// TIA Portal project "Projekt_Serhii_Bodnia" (V19) (continued)

   REGION Timer
       #TP_Remover(IN:= #FlOp_Neg_LS_Auslauf_Band_1.Q,
                   PT:=T#500ms);
       // Störungserkennung: wenn LS_Auslauf länger als 3s aktiv und Band läuft → Stau
       #TON_Störung_LS_Einlauf_Band_0(IN := #LS_Einlauf_Band_0 AND #M_Band_0,
                            PT := T#3s);
       #TON_Störung_LS_Auslauf_Band_0(IN := #LS_Auslauf_Band_0 AND #M_Band_0,
                            PT := T#3s);
       #TON_Störung_LS_Einlauf_Band_1(IN := #LS_Einlauf_Band_1 AND #M_Band_1,
                            PT := T#3s);
       #TON_Störung_LS_Auslauf_Band_1 (IN := #LS_Auslauf_Band_1 AND #M_Band_1,
                            PT := T#3s);
       #TON_Störung_LS_Vision_Sensor (IN := #LS_Vision_Sensor AND #M_Band_0,
                            PT := T#3s);
       #TON_Störung_LS_Arm_0 (IN := #LS_Arm_0 AND #M_Band_0,
                            PT := T#3s);

   END_REGION

    REGION Produktarten
    // Produktart-Rezeptur-Mapping: HMI-Produktauswahl auf Farbewert umrechnen
       IF #Produktart_Linie_0 = 4 THEN
           #Rezeptur_Art_0 := 5;
       ELSIF #Produktart_Linie_0 = 2 THEN
           #Rezeptur_Art_0 := 6;
       END_IF;
       IF #Produktart_Linie_1 = 1 THEN
           #Rezeptur_Art_1 := 2;
       ELSIF #Produktart_Linie_1 = 2 THEN
           #Rezeptur_Art_1 := 1;
       END_IF;
   END_REGION

   REGION Meldungen
       // Störungserkennung: wenn LS_Einlauf oder LS_Auslauf länger als 3s aktiv und Band läuft → Stau
       IF ((#Teil_auf_Band_0 > 5 OR #TON_Störung_LS_Einlauf_Band_0.Q OR #TON_Störung_LS_Auslauf_Band_0.Q
           OR #TON_Störung_LS_Vision_Sensor.Q OR #TON_Störung_LS_Arm_0.Q) AND #M_Band_0 AND NOT #Stop_Modus)
           OR ((#Teil_auf_Band_1 > 5 OR #TON_Störung_LS_Einlauf_Band_1.Q OR #TON_Störung_LS_Auslauf_Band_1.Q) AND #M_Band_1 AND NOT #Stop_Modus) THEN
           // Störungsmerker setzen
           #M_Störung := TRUE;
       END_IF;
       // Störung über HMI quittieren: Bit des Quittierungswortes (HMI_Quittierung)
       IF #Quittierung THEN
           #M_Störung := FALSE;
       END_IF;


   END_REGION

   REGION Sortierung
       IF #FlOp_Pos_LS_Arm_0.Q THEN
           //Farbe des ersten  Werkstücks in der Warteschlange prüfen 
           #Current_Art := #Buffer[0];
           // Array verschieben
           FOR #i := 0 TO 4 DO
               #Buffer[#i] := #Buffer[#i + 1];
           END_FOR;
           // Letzten Element nach dem Verschiebung löschen und den Zäler verringern
           #Buffer[5] := 0;
           IF #Count > 0 THEN
               #Count := #Count - 1;
           END_IF;
       END_IF;

       // Ein- und Ausschaltung Arm_0
       IF #Start_Modus AND (#Current_Art = #Rezeptur_Art_0 AND #FlOp_Pos_LS_Arm_0.Q) THEN
           // Sortierarm EIN: wenn erkannte Produktart dem Rezept entspricht
           #M_Arm_turn_0 := TRUE;
           #M_Arm_Band_0 := TRUE;
       END_IF;
       IF #"FlOp_Neg_LS_Auslauf_Band_0 (1)".Q THEN
           // Arm ausschalten: wenn Teil den Auslauf Band 0 verlassen hat
           #M_Arm_turn_0 := FALSE;
           #M_Arm_Band_0 := FALSE;
       END_IF;

   END_REGION

   REGION Eintag in den Puffer

       IF #FlOp_Pos_LS_Vision_Sensor.Q THEN
           // Farbe speichern
           #Buffer[#Count] := #Vision_Sensor;
           // Platz für den nächsten vorbereiten
           #Count := #Count + 1;
       END_IF;
   END_REGION

   REGION Bänder
       REGION Band_0
           REGION Erfassung der Anzahl der Teileauf dem Band_0
               IF #Start_Modus AND NOT #Stop_Modus THEN
                   // Teilezähler Band_0: zählt aktuell transportierte Teile
                   IF #FlOp_Neg_LS_Einlauf_Band_0.Q THEN
                       #Teil_auf_Band_0 := #Teil_auf_Band_0 + 1;
                   END_IF;
                   IF #Teil_auf_Band_0 > 0 AND (#"FlOp_Neg_LS_Auslauf_Band_0 (1)".Q OR #"FlOp_Neg_LS_Auslauf_Band_0 (2)".Q) THEN
                       #Teil_auf_Band_0 := #Teil_auf_Band_0 - 1;
                   END_IF;
               END_IF;
               IF #Not_Aus_Modus OR #M_Störung THEN
                   #Teil_auf_Band_0 := 0;
               END_IF;
           END_REGION
           REGION Band_0 Steuerung
               // Band_0 läuft solange Teile vorhanden oder neu eingetroffen
               IF #Start_Modus AND (#FlOp_Neg_LS_Einlauf_Band_0.Q OR #Teil_auf_Band_0 > 0) THEN
                   #M_Band_0 := True;
               ELSE
                   #M_Band_0 := FALSE;
               END_IF;

           END_REGION
       END_REGION
       REGION Band_1
           REGION Erfassung der Anzahl der Teileauf dem Band_1
               IF #Start_Modus AND NOT #Stop_Modus THEN
                   // Teilezähler Band 1: zählt aktuell transportierte Teile
                   IF #FlOp_Pos_LS_Einlauf_Band_1.Q THEN
                       #Teil_auf_Band_1 := #Teil_auf_Band_1 + 1;
                   END_IF;
                   IF #Teil_auf_Band_1 > 0 AND #FlOp_Neg_LS_Auslauf_Band_1.Q THEN
                       #Teil_auf_Band_1 := #Teil_auf_Band_1 - 1;
                   END_IF;
               END_IF;
               IF #Not_Aus_Modus OR #M_Störung THEN
                   #Teil_auf_Band_1 := 0;
               END_IF;

           END_REGION
           REGION Band_1 Steuerung
               // Band_1 läuft solange Teile vorhanden oder neu eingetroffen
               IF #Start_Modus AND #FlOp_Pos_LS_Einlauf_Band_1.Q OR #Teil_auf_Band_1 > 0 THEN
                   #M_Band_1 := True;
               ELSE
                   #M_Band_1 := FALSE;
              END_IF;
           END_REGION

       END_REGION

   END_REGION

   REGION Actoren
       // Physische Ausgaben: Bänder und Sortierarm (gesperrt bei Stopp-Modus)
       #Band_0 := #M_Band_0 AND NOT #Stop_Modus;
       #Band_1 := #M_Band_1 AND NOT #Stop_Modus;
       #Arm_turn_0 := #M_Arm_turn_0 AND NOT #Stop_Modus;
       #Arm_Band_0 := #M_Arm_Band_0 AND NOT #Stop_Modus;
       #Remover := #TP_Remover.Q;
       // Gesamtanzahl Fertigteile für HMI
       #Anzahl_Kanister := #CTU_Kanister.CV;
       //
       #Störung := #M_Störung;
   END_REGION
END_FUNCTION_BLOCK

FUNCTION_BLOCK "FB_AbfüllmaschineBand_SCL"   // FB7, SCL
{ S7_Optimized_Access := 'TRUE' }
VERSION : 0.1
   VAR_INPUT
      Start_Mode : Bool;
      Stop_Mode : Bool;
      NotAus_Mode : Bool;
      LS_Einlauf : Bool;
      LS_Auslauf : Bool;
      Diff_Sensor_Tank : Bool;
      Dosing_Aktive : Bool;
      Tank_Level_Meter : Real;
      Quittierung : Bool;
   END_VAR
   VAR_OUTPUT
      Einlaufband : Bool;
      Start_Dosierung : Bool;
      Emitter : Bool;
      "Start Button (Light)" : Bool;
      "Stop Button (Light)" : Bool;
      "Stack Light (Green)" : Bool;
      "Stack Light (Red)" : Bool;
      "Stack Light (Yellow)" : Bool;
      Störung : Bool;
   END_VAR
   VAR
      Stat_Trigger_Neg_Dosing_Stand : F_TRIG;
      Stat_Trigger_Neg_LS_Auslauf : F_TRIG;
      TON_weit_500ms : TON_TIME;
      TON_Störung_Einlauf : TON_TIME;
      TON_Störung_Auslauf : TON_TIME;
      TON_Störung_LS_Tank : TON_TIME;
      iSchritt : Int;
      M_Einlaufband : Bool;
      M_Störung : Bool;
   END_VAR
BEGIN

   REGION Flankenabfragen
       // Statement section REGION
       #Stat_Trigger_Neg_Dosing_Stand(CLK := #Dosing_Aktive); // Fallende Flanke: Dosierung beendet
       #Stat_Trigger_Neg_LS_Auslauf(CLK := #LS_Auslauf); // Fallende Flanke: Flasche am Auslauf
   END_REGION

   REGION Timer
       // Störungserkennung: wenn LS_Einlauf oder LS_Auslauf oder LS_Tank länger als 10s aktiv und Band läuft → Stau
       #"TON_Störung_Einlauf"(IN := #LS_Einlauf AND #M_Einlaufband AND NOT #Stop_Mode,
                            PT := T#10s);
     #TON_Störung_Auslauf(IN := #LS_Auslauf AND #M_Einlaufband AND NOT #Stop_Mode,
                            PT := T#10s);
       #TON_Störung_LS_Tank(IN := #Diff_Sensor_Tank AND #M_Einlaufband AND NOT #Stop_Mode,
                            PT := T#10s);
   END_REGION


   REGION Meldungen
       // Störungserkennung: wenn LS_Einlauf oder LS_Auslauf oder LS_Tank länger als 10s aktiv und Band läuft → Stau

       IF #TON_Störung_Einlauf.Q OR #TON_Störung_Auslauf.Q OR #TON_Störung_LS_Tank.Q THEN
           // Störungsmerker setzen
           #M_Störung := TRUE;
       END_IF;
       // Störung über HMI quittieren: Bit des Quittierungswortes (HMI_Quittierung)
       IF #Quittierung THEN
           #M_Störung := FALSE;
       END_IF;

   END_REGION

   REGION Schrittkette
       IF #NotAus_Mode OR #M_Störung THEN
           // Not-Aus: sofortiger Rücksprung in Initialschritt (alle Aktoren werden abgeschaltet)
           #iSchritt := 0;
       END_IF;

       CASE #iSchritt OF
           0:  // Initialschritt: Startbedingungen prüfen
               // Start nur wenn: Startmodus aktiv UND Füllventil geschlossen UND Tank nicht leer
               IF #Start_Mode  AND (#Tank_Level_Meter >= 1) THEN
                   #iSchritt := 1;
               END_IF;
           1: // Emitter EIN: leere Kanister ausgeben; warten bis Kanister erkannt
               IF #LS_Einlauf THEN
                   #iSchritt := 2;
               END_IF;
           2: // Einlaufband EIN: Kanister unter den Dosierkopf transportieren
              // Übergang wenn Diffusionssensor der Kanister unter dem Tank detektiert
               IF #Diff_Sensor_Tank THEN
                   #iSchritt := 3;
               END_IF;
           3: // Einlaufband AUS; Dosierung starten; warten auf fallende Flanke (Dosierung beendet)
               IF #Stat_Trigger_Neg_Dosing_Stand.Q THEN
                   #iSchritt := 4;
               END_IF;
           4: // Einlaufband EIN (mit TON-Nachlauf 500ms): gefüllte Flasche zum Auslauf schieben
              // Übergang bei fallender Flanke: Kanister hat Auslaufsensor verlassen
               IF #Stat_Trigger_Neg_LS_Auslauf.Q THEN
                   #iSchritt := 1;
               END_IF;

           ELSE  // Unbekannter Schritt: Sicherheitshalber Rücksprung
               #iSchritt := 0;
       END_CASE;
   END_REGION
   REGION Actoren
      // 1. Emitter
       #Emitter := (#iSchritt = 1);
       // 2. Einlaufband
       #TON_weit_500ms(IN := (#iSchritt = 4), PT := T#500ms);
       #Einlaufband := ((#iSchritt = 2) OR #TON_weit_500ms.Q) AND NOT #Stop_Mode;
       #M_Einlaufband := ((#iSchritt = 2) OR #TON_weit_500ms.Q) AND NOT #Stop_Mode;
       // 3. Start_Dosierung
       #Start_Dosierung := (#iSchritt = 3) AND NOT #Stop_Mode;
       // 4. Signallleuchten
       #"Start Button (Light)" := #Start_Mode AND NOT #Stop_Mode;
       #"Stack Light (Green)" := #Start_Mode AND NOT #Stop_Mode;
       #"Stop Button (Light)" := #Stop_Mode;
       #"Stack Light (Red)" := #Stop_Mode;
       #"Stack Light (Yellow)" := #NotAus_Mode;
       //
       #Störung := #M_Störung;

   END_REGION
END_FUNCTION_BLOCK

FUNCTION_BLOCK "FB_Band mit Positionierleisten"   // FB8, SCL
{ S7_Optimized_Access := 'TRUE' }
VERSION : 0.1
   VAR_INPUT
      LS_Einlauf : Bool;
      LS_Auslauf : Bool;
      LS_Positionierer : Bool;
      Start_Modus : Bool;
      Stop_Modus : Bool;
      Not_Aus_Modus : Bool;
      Acknowledge : Bool;
      Quittierung : Bool;
   END_VAR
   VAR_OUTPUT
      Band : Bool;
      Positionierer : Bool;
      Ready_To_Send_Teil : Bool;
      Ready_To_Receive_Teil : Bool;
      Störung : Bool;
   END_VAR
   VAR
      FlOp_Pos_LS_Einlauf : R_TRIG;
      FlOp_Neg_LS_Einlauf : F_TRIG;
      FlOp_Neg_LS_Auslauf : F_TRIG;
      Teil_auf_Band : Int;
      M_Band : Bool;
      M_Positionierer : Bool;
      M_Störung : Bool;
      TON_Störung_LS_Einlauf : TON_TIME;
      TON_Störung_LS_Auslauf : TON_TIME;
      TON_Störung_LS_Positionierer : TON_TIME;
   END_VAR
BEGIN
   REGION Flankenabfragen
       // Alle Flanken müssen am Anfang des Bausteins ausgewertet werden
       #FlOp_Pos_LS_Einlauf(CLK := #LS_Einlauf);
       #FlOp_Neg_LS_Einlauf(CLK := #LS_Einlauf);
       #FlOp_Neg_LS_Auslauf(CLK := #LS_Auslauf);
   END_REGION

   REGION Timers
       // Störungserkennung: wenn LS_Einlauf oder LS_Auslauf länger als 10s aktiv und Band läuft → Stau
       #TON_Störung_LS_Einlauf(IN := #LS_Einlauf AND #M_Band AND NOT #Stop_Modus,
                               PT := T#10s);
       #TON_Störung_LS_Auslauf(IN := #LS_Auslauf AND #M_Band AND NOT #Stop_Modus,
                               PT := T#10s);
       #TON_Störung_LS_Positionierer (IN := #LS_Positionierer AND #M_Band AND NOT #Stop_Modus,
                               PT := T#10s);
   END_REGION

   REGION Meldungen
       // Störungserkennung: wenn LS_Einlauf oder LS_Auslauf länger als 10s aktiv und Band läuft → Stau
       IF #Teil_auf_Band > 3 OR #TON_Störung_LS_Einlauf.Q OR #TON_Störung_LS_Auslauf.Q OR #TON_Störung_LS_Positionierer.Q THEN
           // Störungsmerker setzen
           #M_Störung := TRUE;
       END_IF;
       // Störung über HMI quittieren: Bit des Quittierungswortes (HMI_Quittierung)
       IF #Quittierung THEN
           #M_Störung := FALSE;
       END_IF;

   END_REGION

   REGION Band
       // Teilezähler: zählt Teile auf dem Band
       IF #Start_Modus AND #FlOp_Neg_LS_Einlauf.Q THEN
           // Neues Teil aufgenommen
           #Teil_auf_Band := #Teil_auf_Band + 1;
       END_IF;
       IF #Start_Modus AND #Acknowledge AND #Teil_auf_Band > 0 THEN
           // Teil wurde abgenommen 
           #Teil_auf_Band := #Teil_auf_Band - 1;
       END_IF;
       IF #Not_Aus_Modus THEN
           // Not-Aus: Zähler löschen
           #Teil_auf_Band := 0;
       END_IF;

       // Bandsteuerung: Band einschalten bei steigender Einlaufflanke oder noch Teile vorhanden
       IF #Start_Modus AND #FlOp_Pos_LS_Einlauf.Q OR
           (#LS_Einlauf AND #Teil_auf_Band =0) THEN
           #M_Band := TRUE;
       END_IF;
       IF  #Start_Modus AND #FlOp_Neg_LS_Auslauf.Q THEN
           // Band abschalten sobald Teil das Band verlassen hat
           #M_Band := FALSE;
       END_IF;

   END_REGION

   REGION Positionierer
       // Positionierer klemmt Teil fest zur genauen Ablage durch Pick & Place
       IF #Start_Modus AND NOT #Stop_Modus THEN
           IF #FlOp_Neg_LS_Auslauf.Q THEN
               // Teil hat Auslauf erreicht: klemmen
               #M_Positionierer := TRUE;
           END_IF;
           IF #LS_Positionierer THEN
               // Positionierer vollständig eingeklemmt: fertig
               #M_Positionierer:= FALSE;
           END_IF;
       END_IF;
   END_REGION

   REGION Ready_To_Send & Ready_To_Receive
       IF #Start_Modus AND #LS_Positionierer THEN
           // Weitergabesignal: Teil ist positioniert und bereit für Pick & Place
               #Ready_To_Send_Teil := TRUE;
       END_IF;
       IF #Acknowledge OR #Not_Aus_Modus THEN
           // Pick & Place hat Teil übernommen
           // Ready_To_Send_Teil wird bei Not-Aus zurückgesetzt
               #Ready_To_Send_Teil := FALSE;
       END_IF;

       IF #Teil_auf_Band = 0 THEN
           // Empfangsbereitschaft: Band kann neues Teil aufnehmen wenn es leer ist
           #Ready_To_Receive_Teil := TRUE;
       ELSE
           #Ready_To_Receive_Teil := FALSE;
       END_IF;


   END_REGION

   REGION Actoren
       // Physische Ausgaben: Band und Positionierer werden im Stopp-Modus gesperrt
       #Band := #M_Band AND NOT #Stop_Modus;
       #Positionierer := #M_Positionierer AND NOT #Stop_Modus;
       //
       #Störung := #M_Störung;
   END_REGION
END_FUNCTION_BLOCK

FUNCTION_BLOCK "FB_Palette_Linie"   // FB9, SCL
{ S7_Optimized_Access := 'TRUE' }
VERSION : 0.1
   VAR_INPUT
      LS_Roller_1_Ende : Bool;
      LS_Roller_2_Ende : Bool;
      LS_Roller_3_Beladung : Bool;
      "LS_Roller_3 Ende" : Bool;
      LS_Roller_4_Ende : Bool;
      Start_Modus : Bool;
      Stop_Modus : Bool;
      Not_Aus_Modus : Bool;
      Palette_voll : Bool;
   END_VAR
   VAR_OUTPUT
      Emitter : Bool;
      Roller_Conveyor_1 : Bool;
      Roller_Conveyor_2 : Bool;
      Roller_Conveyor_3 : Bool;
      Roller_Conveyor_4 : Bool;
      Ready_To_Receive_Teil : Bool;
      Remover : Bool;
      Rundumlsmpe : Bool;
      Anzahl_Paletten : Int;
   END_VAR
   VAR
      FlOp_Pos_Emitter : R_TRIG;
      FlOp_Pos_Emitter_1 : R_TRIG;
      FlOp_Neg_LS_Roller_3_Beladung : F_TRIG;
      FlOp_Pos_LS_Roller_1_Ende : R_TRIG;
      FlOp_Pos_LS_Roller_2_Ende : R_TRIG;
      FlOp_Neg_LS_Roller_2_Ende : F_TRIG;
      FlOp_Pos_LS_Roller_4_Ende : R_TRIG;
      FlOp_Neg_LS_Roller_4_Ende : F_TRIG;
      FlOp_Pos_LS_Roller_3_Ende : R_TRIG;
      FlOp_Neg_LS_Roller_3_Ende : F_TRIG;
      TP_Remover : TP_TIME;
      M_Roller_1 : Bool;
      M_Roller_2 : Bool;
      M_Roller_3 : Bool;
      M_Roller_4 : Bool;
      M_nächster_Roller_belegt : Bool;
      M_Ready_To_Receive_Teil : Bool;
      Palette_auf_Roller : Int;
      CTU_Paletten : CTU_INT;
   END_VAR
BEGIN

   REGION Flankenabfragen
       // Emitter-Trigger: neue Palette ausgeben
       // Zwei Trigger-Bedingungen: Sensor 3 aktiv im Start ODER Sensor 2 aktiv und Sensor 3 frei
       #FlOp_Pos_Emitter(CLK := #LS_Roller_3_Beladung AND #Start_Modus);
       #FlOp_Pos_Emitter_1(CLK := #Start_Modus AND #LS_Roller_2_Ende AND NOT #LS_Roller_3_Beladung);
       // Rollenbahn-Sensorflanken
       #FlOp_Pos_LS_Roller_1_Ende(CLK := #LS_Roller_1_Ende);
       #FlOp_Pos_LS_Roller_2_Ende(CLK := #LS_Roller_2_Ende);
       #FlOp_Neg_LS_Roller_2_Ende(CLK := #LS_Roller_2_Ende);
       #FlOp_Pos_LS_Roller_3_Ende(CLK := #"LS_Roller_3 Ende");
       #FlOp_Neg_LS_Roller_3_Ende(CLK := #"LS_Roller_3 Ende");
       #FlOp_Neg_LS_Roller_3_Beladung(CLK := #LS_Roller_3_Beladung);
       #FlOp_Pos_LS_Roller_4_Ende(CLK := #LS_Roller_4_Ende);
       #FlOp_Neg_LS_Roller_4_Ende(CLK := #LS_Roller_4_Ende);

   END_REGION

   REGION Zähler
       // Palettenzähler: Inkrementierung wenn vollbeladene Palette Roller 4 verlässt
       #CTU_Paletten(CU:=#FlOp_Neg_LS_Roller_4_Ende.Q,
                     R:= "FirstScan" OR #Not_Aus_Modus,
                     PV:=0);
   END_REGION

   REGION Timer
       // TP-Impuls für Remover: 2 Sekunden aktiv wenn Palette Roller 4 verlässt
       #TP_Remover(IN := #FlOp_Neg_LS_Roller_4_Ende.Q,
                   PT := T#2s);
   END_REGION

   REGION Ready_To_Send & Ready_To_Receive
       // Beladungsbereitschaft: Palettierbereich ist bereit für neues Teil
       IF #FlOp_Neg_LS_Roller_3_Beladung.Q AND NOT #Palette_voll THEN
           #M_Ready_To_Receive_Teil := TRUE;
       ELSIF #Palette_voll THEN
           // Palette voll: keine weiteren Teile
           #M_Ready_To_Receive_Teil := FALSE;
       END_IF;
   END_REGION

   REGION Roller_1
       // Roller 1: Palette aus Magazin herausführen
       IF #Start_Modus AND (#FlOp_Pos_Emitter.Q OR #FlOp_Pos_Emitter_1.Q) THEN
           // Emitter-Signal: Palette freigeben
           #M_Roller_1 := TRUE;
       END_IF;
       IF #FlOp_Pos_LS_Roller_1_Ende.Q OR #Not_Aus_Modus THEN
           // Palette am Ende von Roller 1 angekommen oder Not-Aus
           #M_Roller_1 := FALSE;
       END_IF;
   END_REGION

   REGION Roller_2
       // Roller 2: Palette von Roller 1 zu Roller 3 (Beladeposition) transportieren
       IF #Start_Modus AND #FlOp_Pos_LS_Roller_1_Ende.Q THEN
           // Palette von Roller 1 übernehmen
           #M_Roller_2 := TRUE;
       END_IF;
       IF #FlOp_Pos_LS_Roller_2_Ende.Q OR #Not_Aus_Modus THEN
           // Palette am Ende von Roller 2 angekommen
           #M_Roller_2 := FALSE;
       END_IF;
       IF NOT #LS_Roller_2_Ende AND #M_Ready_To_Receive_Teil THEN
           #M_nächster_Roller_belegt := TRUE;
       ELSE
           #M_nächster_Roller_belegt := FALSE;
       END_IF;


   END_REGION

   REGION Roller_3
       //Erfassung der Anzahl der Palette auf dem Roller
       IF #Start_Modus  AND #FlOp_Pos_LS_Roller_2_Ende.Q THEN
           #Palette_auf_Roller := #Palette_auf_Roller + 1;
       END_IF;

       IF #Start_Modus AND #FlOp_Pos_LS_Roller_3_Ende.Q AND #Palette_auf_Roller > 0 THEN
           #Palette_auf_Roller := #Palette_auf_Roller - 1;
       END_IF;

       IF #Not_Aus_Modus THEN
           #Palette_auf_Roller := 0;
       END_IF;

       // Steuerung des Roller_3
       IF #Start_Modus AND #FlOp_Neg_LS_Roller_2_Ende.Q AND NOT #M_Ready_To_Receive_Teil THEN
           #M_Roller_3 := TRUE;
       END_IF;
       IF #FlOp_Neg_LS_Roller_3_Beladung.Q THEN
           #M_Roller_3 := FALSE;
       END_IF;
       IF NOT #LS_Roller_3_Beladung AND #Palette_voll THEN
           #M_Roller_3 := TRUE;
       END_IF;
       IF #FlOp_Pos_LS_Roller_3_Ende.Q AND #Palette_auf_Roller = 0 OR #Not_Aus_Modus THEN
           #M_Roller_3 := FALSE;
       END_IF;

   END_REGION

   REGION Roller_4
       // Roller 4: vollbeladene Palette zur Ausgabe transportieren
       IF #Start_Modus AND #FlOp_Neg_LS_Roller_3_Ende.Q THEN
           #M_Roller_4 := TRUE;
       END_IF;
       IF #FlOp_Pos_LS_Roller_4_Ende.Q OR #Not_Aus_Modus THEN
           #M_Roller_4 := FALSE;
       END_IF;

   END_REGION

   REGION Actoren
       // Physische Ausgaben
       // // Bereitschaftssignal für Pick & Place
       #Ready_To_Receive_Teil := #M_Ready_To_Receive_Teil;
       // Palettenausgabe
       #Emitter := #FlOp_Pos_Emitter.Q OR #FlOp_Pos_Emitter_1.Q;
       // 2s-Impuls nach Palettenabgabe
       #Remover := #Start_Modus AND #TP_Remover.Q;
       // Rollenbahnen
       #Roller_Conveyor_1 :=  #M_Roller_1 AND NOT #Stop_Modus;
       #Roller_Conveyor_2 := #M_Roller_2 AND NOT #M_nächster_Roller_belegt AND NOT #Stop_Modus;
       #Roller_Conveyor_3 := #M_Roller_3 AND NOT #Stop_Modus;
       #Roller_Conveyor_4 := #M_Roller_4 AND NOT #Stop_Modus;
       // Gesamtzahl ausgeschleuster Paletten für HMI
       #Anzahl_Paletten := #CTU_Paletten.CV;
   END_REGION
END_FUNCTION_BLOCK

FUNCTION_BLOCK "FB_Pick & Place"   // FB10, SCL
{ S7_Optimized_Access := 'TRUE' }
VERSION : 0.1
   VAR_INPUT
      Sensor_Teil_detect : Bool;
      Start_Modus : Bool;
      Stop_Modus : Bool;
      Not_Aus_Modus : Bool;
      Ready_To_Send_Teil : Bool;
      Ready_To_Receive_Pallet : Bool;
   END_VAR
   VAR_OUTPUT
      X_Set_Point : Real;
      Y_Set_Point : Real;
      Z_Set_Point : Real;
      Grab : Bool;
      Acknowledge_TeIl_Greifen : Bool;
      Pallete_voll : Bool;
      Anzahl_Teil : Int;
      Rundumleuchte : Bool;
   END_VAR
   VAR
      Teil_Position : Array[0..3] of Struct
         X : Real;
         Y : Real;
      END_STRUCT;
      Zähler : Int;
      Schritt : Int;
      "TON_Pick&Place_Schritt_3" : TON_TIME;
      "TON_Pick&Place_Schritt_4" : TON_TIME;
      "TON_Pick&Place_Schritt_5" : TON_TIME;
      "TON_Pick&Place_Schritt_7" : TON_TIME;
      "TON_Pick&Place_Schritt_1" : TON_TIME;
   END_VAR
   VAR RETAIN
      CTU_Teil : CTU_INT;
   END_VAR
   // Teil_Position[0].X := 8.9;
   // Teil_Position[0].Y := 6.4;
   // Teil_Position[1].X := 6.9;
   // Teil_Position[1].Y := 6.4;
   // Teil_Position[2].X := 8.9;
   // Teil_Position[2].Y := 9.5;
   // Teil_Position[3].X := 6.9;
   // Teil_Position[3].Y := 9.5;
BEGIN
   REGION Timer
       // Schritt 1: Wartezeit bis Roboter Greifposition erreicht hat (1500ms)
       #"TON_Pick&Place_Schritt_1"(IN:=#Schritt = 1,
                                   PT:=T#1500ms);
       // Schritt 3: Wartezeit Greifer anheben (1000ms)
       #"TON_Pick&Place_Schritt_3"(IN := #Schritt = 3,
                                   PT := T#1s);
       // Schritt 4: Wartezeit XY-Verfahren zur Zielposition (1500ms)
       #"TON_Pick&Place_Schritt_4"(IN := #Schritt = 4,
                                   PT := T#1500ms);
       // Schritt 5: Wartezeit Greifer absenken (1000ms)
       #"TON_Pick&Place_Schritt_5"(IN := #Schritt = 5,
                                   PT := T#1s);
       // Schritt 7: Wartezeit Greifer nach Ablage anheben (1000ms)
       #"TON_Pick&Place_Schritt_7"(IN := #Schritt = 7,
                                   PT := T#1000ms);
                                END_REGION

   REGION #Zähler
       // Gesamtteilezähler: zählt aufgenommene Teile (steigende Flanke Schritt 3)
       #CTU_Teil(CU:= #Schritt = 3,
                 R:= "FirstScan" OR #Not_Aus_Modus,
                 PV:=0);
       // Ausgabe für HMI-Anzeige
       #Anzahl_Teil := #CTU_Teil.CV;
   END_REGION

   REGION Rundumleuchte
       #Rundumleuchte := #Not_Aus_Modus;
   END_REGION


   CASE #Schritt OF
       0:  // Initialschritt: Roboter in Heimposition (X=0, Y=0, Z=0), 
           #X_Set_Point := 0.0;
           #Y_Set_Point := 0.0;
           #Z_Set_Point := 0.0;
           #Pallete_voll := FALSE;
           IF #Start_Modus THEN
               #Schritt := 1;
           END_IF;
       1:  // Roboter zur Greifposition verfahren (X=0.9, Y=9.5, Z bleibt oben)
           #X_Set_Point := 0.9;
           #Y_Set_Point := 9.5;
           IF #Zähler = 0 THEN
               #Pallete_voll := FALSE;
           END_IF;
           IF #Ready_To_Receive_Pallet AND #Ready_To_Send_Teil AND #"TON_Pick&Place_Schritt_1".Q THEN
               #Schritt := 2;
           END_IF;
       2: // Greifer absenken auf Greiflevel (Z=8.7), auf Teildetektierung warten
               #Z_Set_Point := 8.7;
           IF #Sensor_Teil_detect THEN
               #Grab := TRUE;
               // Quittierung an vorgelagertes Band
               #Acknowledge_TeIl_Greifen := TRUE;
               #Schritt := 3;
           END_IF;
       3: // Greifer anheben mit Teil (Z=0), Quittierung zurücksetzen, Verfahrzeit abwarten
           #Z_Set_Point := 0.0;
           // Quittierung zurücksetzen (Einmalig)
           #Acknowledge_TeIl_Greifen := FALSE;
           IF #"TON_Pick&Place_Schritt_3".Q THEN
               #Schritt := 4;
           END_IF;
       4: // XY-Verfahren zur Ablageposition auf Palette (aus Teil_Position-Array)
          // Zähler bestimmt die aktuelle Ablageposition (0–3, insgesamt 4 Positionen)
           #X_Set_Point := #Teil_Position[#Zähler].X;
           #Y_Set_Point := #Teil_Position[#Zähler].Y;
           IF #"TON_Pick&Place_Schritt_4".Q THEN
               #Schritt := 5;
           END_IF;
       5: // Greifer zur Ablageposition absenken (Z=8.7), Verfahrzeit abwarten
           #Z_Set_Point := 8.7;
           IF #"TON_Pick&Place_Schritt_5".Q THEN
               #Schritt := 6; 
           END_IF;
       6: // Teil ablegen: Greifer öffnen, sofort weiter zu Schritt 7
           #Grab := FALSE;
           #Schritt := 7;
       7: // Greifer nach Ablage anheben, Zähler inkrementieren, zurück zur Greifposition
           #Z_Set_Point := 0.0;
           IF #"TON_Pick&Place_Schritt_7".Q THEN
               // Nächste Ablageposition
               #Zähler := #Zähler + 1;
               #Schritt := 1;
           END_IF;
           // Palette voll nach 4 Teilen (Positionen 0–3): Palette ausschleusen
           IF #Zähler >= 4 THEN
               // Zähler für neue Palette zurücksetzen
               #Zähler := 0;
               // Signal: Palette vollständig beladen
               #Pallete_voll := TRUE;
           END_IF;
       ELSE  // Unbekannter Schritt: bei Not-Aus Rücksprung in Initialschritt
           IF #Not_Aus_Modus THEN
               #Schritt := 0;
           END_IF;

   END_CASE;
END_FUNCTION_BLOCK

FUNCTION_BLOCK "FB_Mode_Manager"   // FB11, SCL
{ S7_Optimized_Access := 'TRUE' }
VERSION : 0.1
   VAR_INPUT
      Start_Taster_Linie_0 : Bool;
      Start_Taster_Linie_1 : Bool;
      Stop_Taster_Linie_0 : Bool;
      Stop_Taster_Linie_1 : Bool;
      Stop_Hauptleitung : Bool;
      NotAus : Bool;
      Rezept_Linie_0 : Real;
      Rezept_Linie_1 : Real;
      Meldung_Störung : Int;
      Quittierung_Störung : Int;
   END_VAR
   VAR_OUTPUT
      Start_Modus_Hauptleitung : Bool;
      Start_Modus_Linie_0 : Bool;
      Start_Modus_Linie_1 : Bool;
      Not_Aus_Modus : Bool;
      Stop_Modus_Hauptleitung : Bool;
      Stop_Modus_Linie_0 : Bool;
      Stop_Modus_Linie_1 : Bool;
   END_VAR
   VAR
      M_Start_Linie_0 : Bool;
      M_Start_Linie_1 : Bool;
      M_Stop_Linie_0 : Bool;
      M_Stop_Linie_1 : Bool;
   END_VAR
BEGIN
   REGION Startmodus
       // Starttaster Linie 0: Betrieb wird nur gestartet, wenn ein gültiges Rezept vorliegt (Rezept <> 0)
       IF #Start_Taster_Linie_0 AND #Rezept_Linie_0 <> 0 THEN
           #M_Start_Linie_0 := TRUE;
           #Start_Modus_Linie_0 := #M_Start_Linie_0;
       END_IF;
       // Starttaster Linie 1: analog zu Linie 0
       IF #Start_Taster_Linie_1 AND #Rezept_Linie_1 <> 0 THEN
           #M_Start_Linie_1 := True;
           #Start_Modus_Linie_1 := #M_Start_Linie_1;
       END_IF;
       // Hauptleitung läuft, sobald mindestens eine Linie im Startmodus ist
       #Start_Modus_Hauptleitung := #M_Start_Linie_0 OR #M_Start_Linie_1;
   END_REGION

   REGION Stopmodus
       // Stopmodus Linie 0: Stopp-Taster setzt, Start-Taster rücksetzt das Halteglied
       IF #"Stop_Taster_Linie_0" OR #Meldung_Störung <> 0 OR #Stop_Hauptleitung THEN
           #M_Stop_Linie_0 := TRUE;
       ELSIF
           #Start_Taster_Linie_0 AND (#Meldung_Störung = 0 OR #Quittierung_Störung <> 0) THEN
           #M_Stop_Linie_0 := FALSE;
       END_IF;
       #Stop_Modus_Linie_0 := #M_Stop_Linie_0;
       // Stopmodus Linie 1: analog zu Linie 0
       IF #"Stop_Taster_Linie_1" OR #Meldung_Störung <> 0 OR #Stop_Hauptleitung THEN
           #M_Stop_Linie_1 := TRUE;
       ELSIF
           #Start_Taster_Linie_1 AND (#Meldung_Störung = 0 OR #Quittierung_Störung <> 0) THEN
           #M_Stop_Linie_1 := FALSE;
       END_IF;
       #Stop_Modus_Linie_1 := #M_Stop_Linie_1;
       // Hauptleitung-Stopp: wenn beide Linien gestoppt sind ODER direkter Hauptleitungsstopp
       IF (#M_Stop_Linie_0 AND #M_Stop_Linie_1) OR #Stop_Hauptleitung OR #Meldung_Störung <> 0 THEN
           #Stop_Modus_Hauptleitung := TRUE;
       ELSIF
           (#Start_Taster_Linie_0 OR #Start_Taster_Linie_1) AND (#Meldung_Störung = 0 OR #Quittierung_Störung <> 0) THEN
           // Jeder Starttaster hebt den Hauptleitungsstopp auf
           #Stop_Modus_Hauptleitung := FALSE;
       END_IF;
   END_REGION

       // Not-Aus-Modus direkt aus dem NotAus-Eingang übernehmen
       #Not_Aus_Modus := #NotAus;
       IF #Not_Aus_Modus THEN
       // Bei Not-Aus: alle Betriebs- und Stoppmodi sofort zurücksetzen
           #Stop_Modus_Hauptleitung := FALSE;
           #Stop_Modus_Linie_0 := FALSE;
           #Stop_Modus_Linie_1 := FALSE;
           #M_Stop_Linie_0 := FALSE;
           #M_Stop_Linie_1 := FALSE;

           #Start_Modus_Hauptleitung := FALSE;
           #Start_Modus_Linie_0 := FALSE;
           #Start_Modus_Linie_1 := FALSE;
           #M_Start_Linie_0 := FALSE;
           #M_Start_Linie_1 := FALSE;
       END_IF;
END_FUNCTION_BLOCK

FUNCTION_BLOCK "FB_Transport_T-Band"   // FB12, SCL
{ S7_Optimized_Access := 'TRUE' }
VERSION : 0.1
   VAR_INPUT
      LS_Einlauf_1 : Bool;
      LS_Einlauf_2 : Bool;
      LS_Ausauf : Bool;
      Start_Modus : Bool;
      Stop_Modus : Bool;
      NotAus_Modus : Bool;
      Quittierung : Bool;
   END_VAR
   VAR_OUTPUT
      Band : Bool;
      Störung : Bool;
   END_VAR
   VAR
      FlOp_Pos_LS_Einlauf_1 : R_TRIG;
      FlOp_Pos_LS_Einlauf_2 : R_TRIG;
      FlOp_Neg_LS_Auslauf : F_TRIG;
      FlOp_Pos_LS_Auslauf : R_TRIG;
      Teil_auf_Band : Int;
      M_Band : Bool;
      M_Störung : Bool;
      TON_Störung_LS_Einlauf_1 : TON_TIME;
      TON_Störung_LS_Einlauf_2 : TON_TIME;
      TON_Störung_LS_Ausauf : TON_TIME;
   END_VAR
BEGIN
   REGION Flankenabfragen
       // Alle Flanken müssen am Anfang des Bausteins aktualisiert werden
       #FlOp_Pos_LS_Einlauf_1(CLK := #LS_Einlauf_1);
       #FlOp_Pos_LS_Einlauf_2(CLK := #LS_Einlauf_2);
       #FlOp_Neg_LS_Auslauf(CLK := #LS_Ausauf);
       #FlOp_Pos_LS_Auslauf(CLK := #LS_Ausauf);

   END_REGION

   REGION Timers
       #TON_Störung_LS_Einlauf_1 (IN := #LS_Einlauf_1 AND #M_Band AND NOT #Stop_Modus,
                                  PT := T#10s);
       #TON_Störung_LS_Einlauf_2 (IN := #LS_Einlauf_2 AND #M_Band AND NOT #Stop_Modus,
                                  PT := T#10s);
       #TON_Störung_LS_Ausauf(IN := #LS_Ausauf AND #M_Band AND NOT #Stop_Modus,
                            PT := T#10s);
   END_REGION

   REGION Meldungen
       // Störungserkennung: wenn LS_Einlauf oder LS_Auslauf länger als 10s aktiv und Band läuft → Stau
       IF (#Teil_auf_Band > 3 OR #TON_Störung_LS_Einlauf_1.Q OR #TON_Störung_LS_Einlauf_2.Q OR #TON_Störung_LS_Ausauf.Q) AND #M_Band THEN
           // Störungsmerker setzen
           #M_Störung := TRUE;
       END_IF;
       // Störung über HMI quittieren: Bit des Quittierungswortes (HMI_Quittierung)
       IF #Quittierung THEN
           #M_Störung := FALSE;
       END_IF;

   END_REGION

   REGION Erfassung der Anzahl der Teileauf dem Band
       // Teilezähler: Inkrementierung bei jedem neuen Teil von beiden Einläufen
       IF #Start_Modus AND NOT #Stop_Modus AND (#FlOp_Pos_LS_Einlauf_1.Q OR #FlOp_Pos_LS_Einlauf_2.Q) THEN
           #Teil_auf_Band := #Teil_auf_Band + 1;
       END_IF;
       // Dekrementierung wenn Teil den Auslauf verlässt
       IF #Start_Modus AND NOT #Stop_Modus AND #FlOp_Neg_LS_Auslauf.Q AND #Teil_auf_Band > 0 THEN
           #Teil_auf_Band := #Teil_auf_Band - 1;
       END_IF;
       // Not-Aus: Teilezähler zurücksetzen 
       IF #NotAus_Modus THEN
           #Teil_auf_Band := 0;
       END_IF;
   END_REGION

   REGION Band
       // Band läuft nur wenn Teil von Einlauf 1 angekommen ODER noch Teile auf Band
       IF #Start_Modus AND (#FlOp_Pos_LS_Einlauf_1.Q OR #Teil_auf_Band > 0) THEN
           #M_Band := True;
       ELSE
           #M_Band := FALSE;
       END_IF;
       // Not-Aus und Störung: Bandmerker sofort löschen
       IF #NotAus_Modus OR #M_Störung THEN
           #M_Band := FALSE;
       END_IF;

   END_REGION

   REGION Aktoren
       // Physischer Ausgang: Band läuft nur wenn Merker gesetzt UND kein Stopp-Modus
       #Band := #M_Band AND NOT #Stop_Modus;
       #Störung := #M_Störung;
   END_REGION
END_FUNCTION_BLOCK

FUNCTION_BLOCK "FB_Laufzeit"   // FB13, SCL
{ S7_Optimized_Access := 'TRUE' }
VERSION : 0.1
   VAR_INPUT
      Start_Modus : Bool;
      Stop_Modus : Bool;
   END_VAR
   VAR_OUTPUT
      Run_Hours : Int;
      Run_Minutes : Int;
      Run_Sekunden : Int;
   END_VAR
   VAR
      Run_Time_Text : String;
      R_Trig_1s : R_TRIG;
      Seconds_Total : DInt;
   END_VAR
BEGIN
   REGION Flankenabfragen
       // Steigende Flanke des 1-Hz-Systemtakts (Clock_1Hz) zur sekundengenauen Zeitmessung
       #R_Trig_1s(CLK := "Clock_1Hz");
   END_REGION

   IF "FirstScan" OR NOT #Start_Modus THEN
       // Betriebsstundenzähler zurücksetzen beim ersten Aufruf ODER wenn Startmodus inaktiv
       #Seconds_Total := 0;
       #Run_Sekunden := 0;
       #Run_Minutes := 0;
       #Run_Hours := 0;
   END_IF;

   IF #R_Trig_1s.Q AND #Start_Modus AND NOT #Stop_Modus THEN
       // Sekundenzähler inkrementieren: nur wenn Startmodus aktiv UND kein Stopp
       #Seconds_Total := #Seconds_Total +1;
   END_IF;
   // Umrechnung Gesamtsekunden → Stunden, Minuten, Sekunden
   #Run_Sekunden := DINT_TO_INT(#Seconds_Total MOD 60);
   #Run_Minutes := DINT_TO_INT((#Seconds_Total / 60) MOD 60);
   #Run_Hours := DINT_TO_INT(#Seconds_Total / 3600);
END_FUNCTION_BLOCK

FUNCTION "FC_Scalierung" : Void   // FC1, FBD
{ S7_Optimized_Access := 'TRUE' }
VERSION : 0.1
   VAR_INPUT
      Tankfüllvolumen_Rezept_L_0 : Real;
      Tankfüllvolumen_Rezept_L_1 : Real;
      Tank_0_Level_Meter : Real;
      Tank_1_Level_Meter : Real;
      Dosiervolumen_Rezept_0 : Real;
      Dosiervolumen_Rezept_1 : Real;
   END_VAR
   VAR_OUTPUT
      Input_HMI_Level_L_0 : Real;
      Input_HMI_Level_L_1 : Real;
      Tank_0_level : Real;
      Tank_1_level : Real;
      Tankfüllvolumen_L_0 : Real;
      Tankfüllvolumen_L_1 : Real;
      Dosiervolumen_L_0 : Real;
      Dosiervolumen_L_1 : Real;
   END_VAR
   VAR_TEMP
      Input_Level_norm_0 : Real;
      Input_Level_norm_1 : Real;
      Tank_Level_norm_0 : Real;
      Tank_Level_norm_1 : Real;
   END_VAR
BEGIN

REGION Network 1: Input_HMI_Level_0
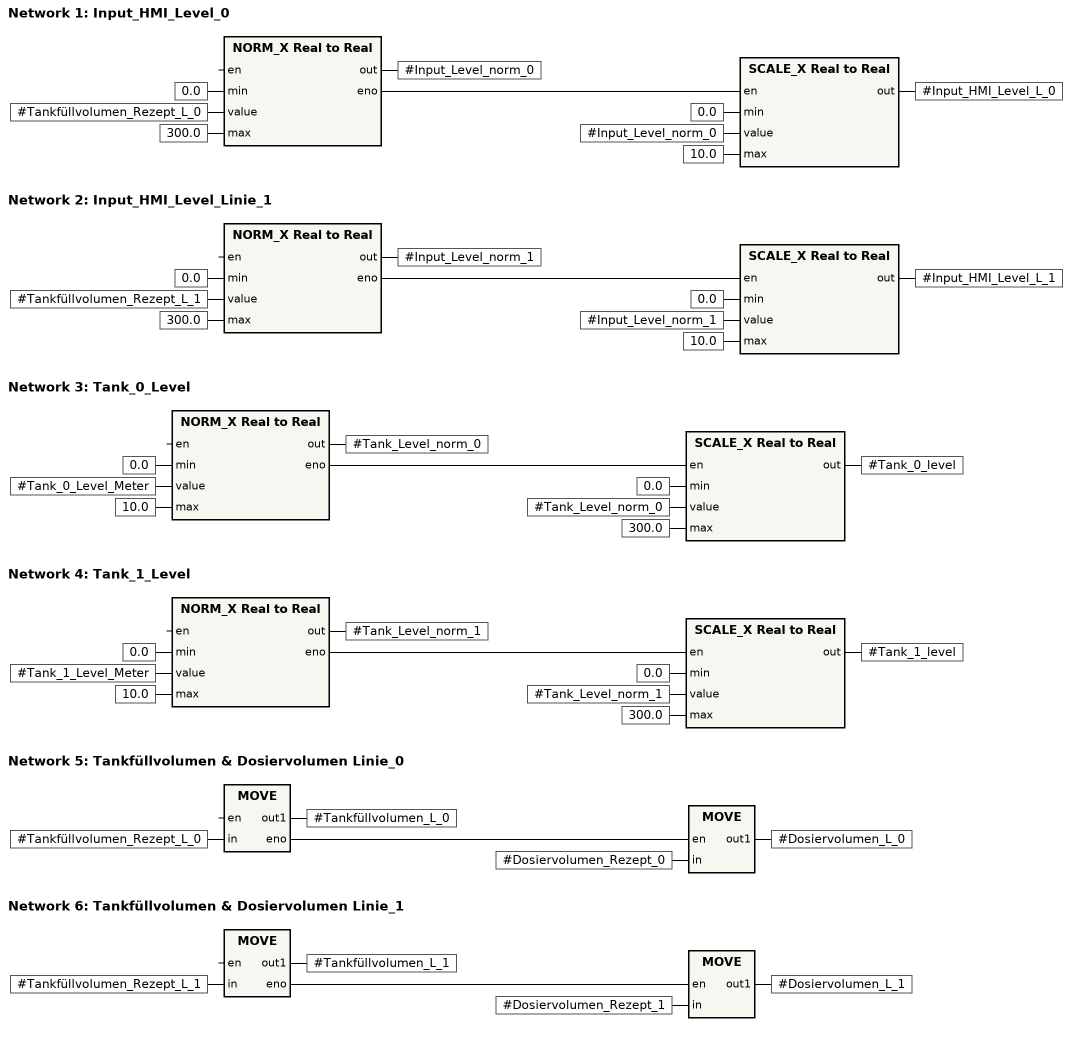
   #Input_Level_norm_0 := NORM_X(MIN := 0.0, VALUE := #Tankfüllvolumen_Rezept_L_0, MAX := 300.0);
   #Input_HMI_Level_L_0 := SCALE_X(MIN := 0.0, VALUE := #Input_Level_norm_0, MAX := 10.0);
END_REGION

REGION Network 2: Input_HMI_Level_Linie_1
   #Input_Level_norm_1 := NORM_X(MIN := 0.0, VALUE := #Tankfüllvolumen_Rezept_L_1, MAX := 300.0);
   #Input_HMI_Level_L_1 := SCALE_X(MIN := 0.0, VALUE := #Input_Level_norm_1, MAX := 10.0);
END_REGION

REGION Network 3: Tank_0_Level
   #Tank_Level_norm_0 := NORM_X(MIN := 0.0, VALUE := #Tank_0_Level_Meter, MAX := 10.0);
   #Tank_0_level := SCALE_X(MIN := 0.0, VALUE := #Tank_Level_norm_0, MAX := 300.0);
END_REGION

REGION Network 4: Tank_1_Level
   #Tank_Level_norm_1 := NORM_X(MIN := 0.0, VALUE := #Tank_1_Level_Meter, MAX := 10.0);
   #Tank_1_level := SCALE_X(MIN := 0.0, VALUE := #Tank_Level_norm_1, MAX := 300.0);
END_REGION

REGION Network 5: Tankfüllvolumen & Dosiervolumen Linie_0
   #Tankfüllvolumen_L_0 := #Tankfüllvolumen_Rezept_L_0;
   #Dosiervolumen_L_0 := #Dosiervolumen_Rezept_0;
END_REGION

REGION Network 6: Tankfüllvolumen & Dosiervolumen Linie_1
   #Tankfüllvolumen_L_1 := #Tankfüllvolumen_Rezept_L_1;
   #Dosiervolumen_L_1 := #Dosiervolumen_Rezept_1;
END_REGION
END_FUNCTION

FUNCTION "MHJ-PLC-Lab-Function-S71200" : Void   // FC9000, SCL
{ S7_Optimized_Access := 'TRUE' }
VERSION : 0.1
   VAR_TEMP
      rdTimeReturn : Int;
      outputTime : DTL;
      SyncVal : Byte;
      forVal : Int;
      forVal_2 : Int;
      Value : Byte;
   END_VAR
   VAR CONSTANT
      CompVal : Byte := 16#34;
      Value_01 : Byte := 16#11;
      Value_01_DW : DWord := 16#A165_D992;
      Value_02_DW : DWord := 16#58BE_4401;
   END_VAR
BEGIN

   #Value:=PEEK(area := 16#82,
        dbNumber := 0,
        byteOffset := 511);
   #Value := #Value + 1;

   POKE(area := 16#82,
        dbNumber := 0,
        byteOffset := 511,
        value := #Value);

   POKE(area:=16#81,
        dbNumber:=0,
        byteOffset:=1016,
        value:=#Value_01_DW);
   POKE(area := 16#81,
        dbNumber := 0,
        byteOffset := 1020,
        value := #Value_02_DW);

   POKE(area := 16#81,
        dbNumber := 0,
        byteOffset := 511,
        value := B#16#00);